// TIA Portal project "Project_python" (V16)

(* hardware
DEVICE "S7-1200 station_2"  S7-1200 Station
   slot 0: "Rack_0"  S7-1200 Rack  Rack  V1.0
   slot 1: "PLC_2"  CPU 1215C DC/DC/DC  6ES7 215-1AG40-0XB0  V4.4
*)

// ===== PLC "PLC_2"  CPU 1215C DC/DC/DC =====

VAR_GLOBAL   // PLC tag table "Default tag table"
   "LIGA" AT %M0.0 : Bool;
   "DESLIGA" AT %M0.1 : Bool;
   "MOTOR" AT %M0.2 : Bool;
   "MEMORIA_SINT" AT %MB10 : SInt;
   "LIGA_IO" AT %I0.0 : Bool;
   "DESLIGA_IO" AT %I0.1 : Bool;
   "MOTOR_IO" AT %Q0.0 : Bool;
   "MEMORIA_INT" AT %MW14 : Int;
   "MEMORIA_DINT" AT %MD16 : DInt;
   "MEMORIA_REAL" AT %MD20 : Real;
   "MOTOR2" AT %M0.3 : Bool;
   "MOTOR3" AT %M0.4 : Bool;
END_VAR

DATA_BLOCK "BASE"   // DB120
{ S7_Optimized_Access := 'FALSE' }
VERSION : 0.1
   VAR
      LIGA_DB : Bool;
      DESLIGA_DB : Bool;
      MOTOR_DB : Bool;
      CONTADOR : IEC_UCOUNTER;
      CONTAGEM_LIGADO : UInt;
      CONTAGEM_DESLIGADO : UInt;
      TEMPORIZADOR : IEC_TIMER;
   END_VAR
BEGIN
END_DATA_BLOCK

// folder: System blocks/Program resources

DATA_BLOCK "CONTADOR_SISTEMA"   // DB1
{ S7_Optimized_Access := 'TRUE' }
AUTHOR : Simatic
FAMILY : IEC
NAME : UCNTR
VERSION : 1.2
// stored: InstanceOfName IEC_UCOUNTER
"IEC_UCOUNTER"
BEGIN
END_DATA_BLOCK

DATA_BLOCK "TEMPORIZADOR_SISTEMA"   // DB2
{ S7_Optimized_Access := 'TRUE' }
AUTHOR : Simatic
FAMILY : IEC
NAME : IEC_TMR
VERSION : 1.0
// stored: InstanceOfName IEC_TIMER
"IEC_TIMER"
BEGIN
END_DATA_BLOCK

// folder: (top level)

ORGANIZATION_BLOCK "Main"   // OB1, LAD, ProgramCycle
TITLE = "Main Program Sweep (Cycle)"
{ S7_Optimized_Access := 'TRUE' }
VERSION : 0.1
   VAR_INPUT
      Initial_Call : Bool;   // Initial call of this OB
      Remanence : Bool;   // =True, if remanent data are available
   END_VAR
BEGIN

REGION Network 1
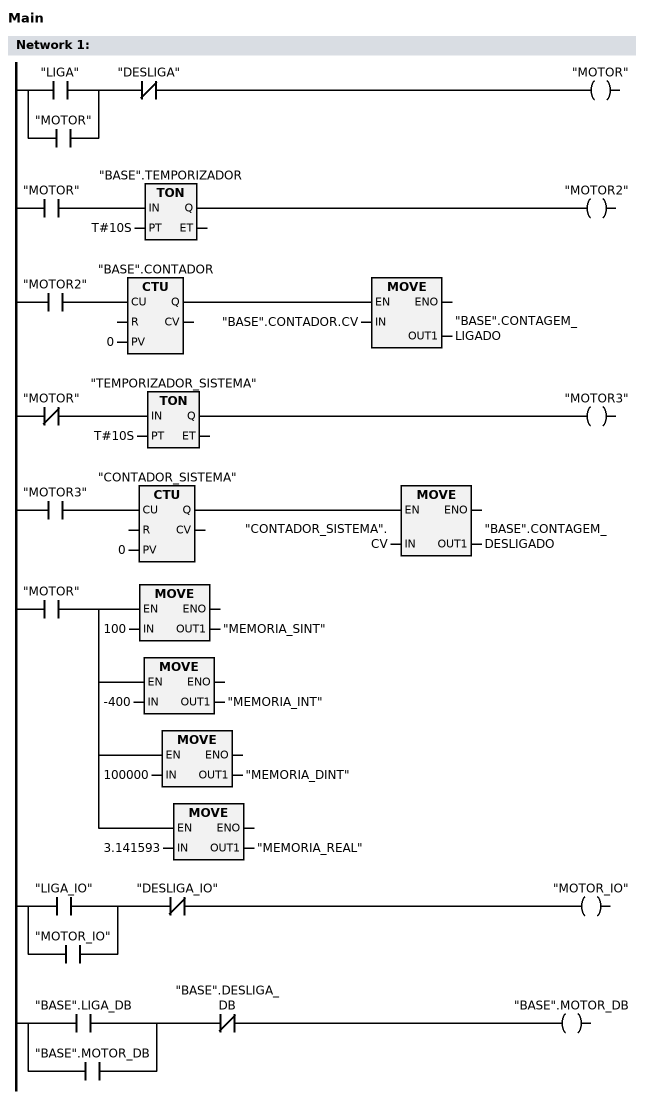
   "MOTOR" := ("LIGA" OR "MOTOR") AND NOT "DESLIGA";
   "BASE".TEMPORIZADOR.TON(IN := "MOTOR", PT := T#10S);
   "MOTOR2" := "BASE".TEMPORIZADOR.Q;
   "BASE".CONTADOR.CTU(CU := "MOTOR2", PV := 0);
   IF "BASE".CONTADOR.Q THEN "BASE".CONTAGEM_LIGADO := "BASE".CONTADOR.CV; END_IF;
   "TEMPORIZADOR_SISTEMA".TON(IN := NOT "MOTOR", PT := T#10S);
   "MOTOR3" := "TEMPORIZADOR_SISTEMA".Q;
   "CONTADOR_SISTEMA".CTU(CU := "MOTOR3", PV := 0);
   IF "CONTADOR_SISTEMA".Q THEN "BASE".CONTAGEM_DESLIGADO := "CONTADOR_SISTEMA".CV; END_IF;
   IF "MOTOR" THEN
       "MEMORIA_SINT" := 100;
       "MEMORIA_INT" := -400;
       "MEMORIA_DINT" := 100000;
       "MEMORIA_REAL" := 3.141593;
   END_IF;
   "MOTOR_IO" := ("LIGA_IO" OR "MOTOR_IO") AND NOT "DESLIGA_IO";
   "BASE".MOTOR_DB := ("BASE".LIGA_DB OR "BASE".MOTOR_DB) AND NOT "BASE".DESLIGA_DB;
END_REGION
END_ORGANIZATION_BLOCK